   Line "Line_420" at 976,739 size 25x0
      Appearance <- "step_vessel_5"
      Visibility <- "step_vessel_5_proses"
   Line "Line_421" at 748,400 size 25x11
      Appearance <- "step_vessel_4"
      Visibility <- "step_vessel_4_proses"
   Line "Line_422" at 752,412 size 36x78
      Appearance <- "step_vessel_4"
      Visibility <- "step_vessel_4_proses"
   Line "Line_423" at 788,488 size 0x11
      Appearance <- "step_vessel_4"
      Visibility <- "step_vessel_4_proses"
   Line "Line_426" at 767,595 size 21x144
      Appearance <- "step_vessel_4"
      Visibility <- "step_vessel_4_proses"
   Line "Line_427" at 788,579 size 0x19
      Appearance <- "step_vessel_4"
      Visibility <- "step_vessel_4_proses"
   Line "Line_428" at 764,739 size 25x0
      Appearance <- "step_vessel_4"
      Visibility <- "step_vessel_4_proses"
   Line "Line_429" at 536,400 size 25x11
      Appearance <- "step_vessel_3"
   Line "Line_430" at 540,412 size 36x78
      Appearance <- "step_vessel_3"
   Line "Line_431" at 576,488 size 0x11
      Appearance <- "step_vessel_3"
   Line "Line_432" at 748,400 size 25x11
      Appearance <- "step_vessel_4"
   Line "Line_433" at 752,412 size 36x78
      Appearance <- "step_vessel_4"
   Line "Line_434" at 788,488 size 0x11
      Appearance <- "step_vessel_4"
   Line "Line_435" at 960,400 size 25x11
      Appearance <- "step_vessel_5"
   Line "Line_436" at 964,412 size 36x78
      Appearance <- "step_vessel_5"
   Line "Line_437" at 1000,488 size 0x11
      Appearance <- "step_vessel_5"
   Line "Line_438" at 1172,400 size 25x11
      Appearance <- "step_vessel_6"
   Line "Line_439" at 1176,412 size 36x78
      Appearance <- "step_vessel_6"
   Line "Line_440" at 1212,488 size 0x11
      Appearance <- "step_vessel_6"
   Line "Line_441" at 1384,400 size 25x11
      Appearance <- "step_vessel_7"
   Line "Line_442" at 1388,412 size 36x78
      Appearance <- "step_vessel_7"
   Line "Line_443" at 1424,488 size 0x11
      Appearance <- "step_vessel_7"
   Line "Line_450" at 555,595 size 21x144
      Appearance <- "step_vessel_3"
   Line "Line_451" at 576,579 size 0x19
      Appearance <- "step_vessel_3"
   Line "Line_452" at 552,739 size 25x0
      Appearance <- "step_vessel_3"
   Line "Line_453" at 767,595 size 21x144
      Appearance <- "step_vessel_4"
   Line "Line_454" at 788,579 size 0x19
      Appearance <- "step_vessel_4"
   Line "Line_455" at 764,739 size 25x0
      Appearance <- "step_vessel_4"
   Line "Line_457" at 979,595 size 21x144
      Appearance <- "step_vessel_5"
   Line "Line_458" at 1000,579 size 0x19
      Appearance <- "step_vessel_5"
   Line "Line_459" at 976,739 size 25x0
      Appearance <- "step_vessel_5"
   Line "Line_461" at 1191,595 size 21x144
      Appearance <- "step_vessel_6"
   Line "Line_462" at 1212,579 size 0x19
      Appearance <- "step_vessel_6"
   Line "Line_463" at 1188,739 size 25x0
      Appearance <- "step_vessel_6"
   Line "Line_464" at 1403,595 size 21x144
      Appearance <- "step_vessel_7"
   Line "Line_465" at 1424,579 size 0x19
      Appearance <- "step_vessel_7"
   Line "Line_466" at 1400,739 size 25x0
      Appearance <- "step_vessel_7"
   Polygon "Polygon_217" at 123,352 size 58x419
      Appearance <- "ISI TANK 1"
      Visibility <- "ISI TANK 1"
   Line "Line_468" at 124,432 size 57x0
      Visibility <- "ISI TANK 1"
   Line "Line_469" at 142,385 size 21x0
      Visibility <- "ISI TANK 1"
   Line "Line_470" at 124,680 size 56x0
      Visibility <- "ISI TANK 1"
   Polygon "Polygon_218" at 335,352 size 58x419
      Appearance <- "ISI TANK 2"
      Visibility <- "ISI TANK 2"
   Line "Line_471" at 336,432 size 57x0
      Visibility <- "ISI TANK 2"
   Line "Line_472" at 354,385 size 21x0
      Visibility <- "ISI TANK 2"
   Line "Line_473" at 336,680 size 56x0
      Visibility <- "ISI TANK 2"
   Polygon "Polygon_219" at 547,352 size 58x419
      Appearance <- "ISI TANK 3"
      Visibility <- "ISI TANK 3"
   Line "Line_474" at 548,432 size 57x0
      Visibility <- "ISI TANK 3"
   Line "Line_475" at 566,385 size 21x0
      Visibility <- "ISI TANK 3"
   Line "Line_476" at 548,680 size 56x0
      Visibility <- "ISI TANK 3"
   Polygon "Polygon_220" at 759,352 size 58x419
      Appearance <- "ISI TANK 4"
      Visibility <- "ISI TANK 4"
   Line "Line_477" at 760,432 size 57x0
      Visibility <- "ISI TANK 4"
   Line "Line_478" at 778,385 size 21x0
      Visibility <- "ISI TANK 4"
   Line "Line_479" at 760,680 size 56x0
      Visibility <- "ISI TANK 4"
   Polygon "Polygon_221" at 971,352 size 58x419
      Appearance <- "ISI TANK 5"
      Visibility <- "ISI TANK 5"
   Line "Line_480" at 972,432 size 57x0
      Visibility <- "ISI TANK 5"
   Line "Line_481" at 990,385 size 21x0
      Visibility <- "ISI TANK 5"
   Line "Line_482" at 972,680 size 56x0
      Visibility <- "ISI TANK 5"
   Polygon "Polygon_222" at 1183,352 size 58x419
      Appearance <- "ISI TANK 6"
      Visibility <- "ISI TANK 6"
   Line "Line_483" at 1184,432 size 57x0
      Visibility <- "ISI TANK 6"
   Line "Line_484" at 1202,385 size 21x0
      Visibility <- "ISI TANK 6"
   Line "Line_485" at 1184,680 size 56x0
      Visibility <- "ISI TANK 6"
   Polygon "Polygon_223" at 1395,352 size 58x419
      Appearance <- "ISI TANK 7"
      Visibility <- "ISI TANK 7"
   Line "Line_486" at 1396,432 size 57x0
      Visibility <- "ISI TANK 7"
   Line "Line_487" at 1414,385 size 21x0
      Visibility <- "ISI TANK 7"
   Line "Line_488" at 1396,680 size 56x0
      Visibility <- "ISI TANK 7"
   Line "Line_489" at 105,898 size 0x48
      Visibility <- "step_vessel_1_proses"
      Appearance <- "step_vessel_1_proses"
   Line "Line_490" at 102,948 size 40x0
      Appearance <- "step_vessel_1_proses"
      Visibility <- "step_vessel_1_proses"
   Rectangle "Rectangle_10" at 75,874 size 1423x33
      Appearance <- "step_vessel_1_proses"
      Visibility <- "step_vessel_1_proses"
   Line "Line_491" at 105,898 size 0x48
      Appearance <- "step_vessel_2_proses"
      Visibility <- "step_vessel_2_proses"
   Line "Line_492" at 102,948 size 40x0
      Appearance <- "step_vessel_2_proses"
      Visibility <- "step_vessel_2_proses"
   Rectangle "Rectangle_11" at 75,874 size 1423x33
      Visibility <- "step_vessel_2_proses"
      Appearance <- "step_vessel_2_proses"
   Line "Line_493" at 105,898 size 0x48
      Appearance <- "step_vessel_3_proses"
      Visibility <- "step_vessel_3_proses"
   Line "Line_494" at 102,948 size 40x0
      Appearance <- "step_vessel_3_proses"
      Visibility <- "step_vessel_3_proses"
   Rectangle "Rectangle_12" at 75,874 size 1423x33
      Appearance <- "step_vessel_3_proses"
      Visibility <- "step_vessel_3_proses"
   Group "proses_3" at 75,874 size 1423x74
   Line "Line_495" at 105,898 size 0x48
      Appearance <- "step_vessel_4_proses"
      Visibility <- "step_vessel_4_proses"
   Line "Line_496" at 102,948 size 40x0
      Appearance <- "step_vessel_4_proses"
      Visibility <- "step_vessel_4_proses"
   Rectangle "Rectangle_13" at 75,874 size 1423x33
      Appearance <- "step_vessel_4_proses"
      Visibility <- "step_vessel_4_proses"
   Group "proses_4" at 75,874 size 1423x74
   Line "Line_497" at 105,898 size 0x48
      Appearance <- "step_vessel_5_proses"
      Visibility <- "step_vessel_5_proses"
   Line "Line_498" at 102,948 size 40x0
      Appearance <- "step_vessel_5_proses"
      Visibility <- "step_vessel_5_proses"
   Rectangle "Rectangle_14" at 75,874 size 1423x33
      Appearance <- "step_vessel_5_proses"
      Visibility <- "step_vessel_5_proses"
   Group "proses_5" at 75,874 size 1423x74
   Line "Line_499" at 105,898 size 0x48
      Visibility <- "step_vessel_6_proses"
      Appearance <- "step_vessel_6_proses"
   Line "Line_500" at 102,948 size 40x0
      Appearance <- "step_vessel_6_proses"
      Visibility <- "step_vessel_6_proses"
   Rectangle "Rectangle_15" at 75,874 size 1423x33
      Appearance <- "step_vessel_6_proses"
      Visibility <- "step_vessel_6_proses"
   Group "proses_6" at 75,874 size 1423x74
   Line "Line_501" at 105,898 size 0x48
      Visibility <- "step_vessel_7_proses"
      Appearance <- "step_vessel_7_proses"
   Line "Line_502" at 102,948 size 40x0
      Appearance <- "step_vessel_7_proses"
      Visibility <- "step_vessel_7_proses"
   Rectangle "Rectangle_16" at 75,874 size 1423x33
      Visibility <- "step_vessel_7_proses"
      Appearance <- "step_vessel_7_proses"
   Group "proses_7" at 75,874 size 1423x74
   Line "Line_379" at 324,400 size 25x11
      Appearance <- "step_vessel_2"
   Line "Line_380" at 328,412 size 36x78
      Appearance <- "step_vessel_2"
   Line "Line_381" at 364,488 size 0x11
      Appearance <- "step_vessel_2"
   Line "Line_505" at 343,595 size 21x144
      Appearance <- "step_vessel_2"
   Line "Line_506" at 364,579 size 0x19
      Appearance <- "step_vessel_2"
   Line "Line_507" at 340,739 size 25x0
      Appearance <- "step_vessel_2"

screen "storage" 1600x1200
   GraphicView "Graphic view_3" at 191,109 size 312x345; Picture "Graphic_8"
   GraphicView "Graphic view_1" at 191,538 size 312x345; Picture "Graphic_8"
   Group "Group" at 704,26 size 95x303; Picture "Graphic_10"
   Group "Group_2" at 704,453 size 95x303; Picture "Graphic_10"
   Group "Group_3" at 898,453 size 95x303; Picture "Graphic_10"
   Group "Group_4" at 898,26 size 95x303; Picture "Graphic_10"
   GraphicView "Graphic view_45" at 1130,217 size 45x48; Picture "Graphic_56"
   GraphicView "Graphic view_44" at 1130,147 size 47x75; Picture "Graphic_55"
   GraphicView "Graphic view_46" at 1218,217 size 45x48; Picture "Graphic_56"
   GraphicView "Graphic view_47" at 1218,147 size 47x75; Picture "Graphic_55"
   GraphicView "Graphic view_49" at 1130,662 size 45x48; Picture "Graphic_56"
   GraphicView "Graphic view_50" at 1130,592 size 47x75; Picture "Graphic_55"
   GraphicView "Graphic view_51" at 1218,662 size 45x48; Picture "Graphic_56"
   GraphicView "Graphic view_52" at 1218,592 size 47x75; Picture "Graphic_55"
   Button "Button_1" at 633,851 size 192x32; TextOn 'Screen_1'; TextOff 'Vessel'
      on Click: ActivateScreen("vessel", 0)
   Button "Button_2" at 880,851 size 192x32; TextOn 'Screen_3'; TextOff 'Supply'
      on Click: ActivateScreen("supply", 0)
   TextField "Text field_9" at 1484,420 size 16x22; Text 'D'
   IOField "I/O field_25" at 1216,276 size 38x17; FormatPattern 9999999
      Appearance <- "VP FLAVOUR"
   TextField "Text field_13" at 1252,276 size 25x18; Text 'bar'
   IOField "I/O field_26" at 1022,229 size 38x17; FormatPattern 9999999
      Appearance <- "VP FLAVOUR"
   TextField "Text field_14" at 1058,229 size 23x18; Text 'º C'
   IOField "I/O field_1" at 1116,24 size 38x17; FormatPattern 9999999
      Appearance <- "VP FLAVOUR"
   TextField "Text field_10" at 1152,24 size 25x18; Text 'bar'
   IOField "I/O field_2" at 1022,655 size 38x17; FormatPattern 9999999
      Appearance <- "VP HIDROLIC"
   TextField "Text field_1" at 1058,655 size 23x18; Text 'º C'
   IOField "I/O field_3" at 1216,724 size 38x17; FormatPattern 9999999
      Appearance <- "VP HIDROLIC"
   TextField "Text field_5" at 1252,724 size 25x18; Text 'bar'
   IOField "I/O field_4" at 1116,480 size 38x17; FormatPattern 9999999
      Appearance <- "VP HIDROLIC"
   TextField "Text field_4" at 1152,480 size 25x18; Text 'bar'
   IOField "I/O field_5" at 798,711 size 38x17; FormatPattern 9999999
      Appearance <- "VP HIDROLIC"
   TextField "Text field_6" at 834,711 size 23x18; Text 'º C'
   IOField "I/O field_6" at 798,287 size 38x17; FormatPattern 9999999
      Appearance <- "VP FLAVOUR"
   TextField "Text field_7" at 834,287 size 23x18; Text 'º C'
   IOField "I/O field_7" at 614,47 size 38x17; FormatPattern 9999999
      Appearance <- "VP FLAVOUR"
   TextField "Text field_2" at 650,47 size 23x18; Text 'º C'
   IOField "I/O field_8" at 614,471 size 38x17; FormatPattern 9999999
      Appearance <- "VP HIDROLIC"
   TextField "Text field_3" at 650,471 size 23x18; Text 'º C'
   TextField "Text field_8" at 195,529 size 138x23; Text 'TANK HIDROLIK'
   TextField "Text field_12" at 1449,457 size 117x23; Text 'FROM VESSEL'
   GraphicView "Graphic view_4" at 17,916 size 156x94; Picture "Graphic_72"
   GraphicView "Graphic view_7" at 17,481 size 156x94; Picture "Graphic_72"
   Group "Group_10" at 209,458 size 22x12
   Group "Group_1" at 209,890 size 22x12
   Group "Group_6" at 985,57 size 363x395
   Group "Group_8" at 792,83 size 114x184
   Group "Group_11" at 346,86 size 364x39
   Group "Group_12" at 346,86 size 364x39
   Group "Group_13" at 984,507 size 451x318
   Group "Group_15" at 790,516 size 116x179
   Group "Group_17" at 346,513 size 364x42
   Group "Group_18" at 346,513 size 364x42
   Circle "Circle_1" at 320,266 size 43x43
      Appearance <- "tank flavour OK"
   Circle "Circle_2" at 320,698 size 43x43
      Appearance <- "tank hidrolic OK"
   Button "Button_3" at 633,812 size 96x32; TextOff 'Transfer'
      on Press: function_b14e0dd5("transfer", 0)
   Button "Button_4" at 790,810 size 109x34; TextOff 'Auto'; TextList "moded"
      on Click: InvertBit("mode")
      ProcessValue <- "mode"
      Appearance <- "mode"
   Group "Group_19" at 1366,449 size 144x36
   Group "Group_20" at 1366,449 size 144x36
   Group "Group_21" at 1366,449 size 144x36
   Group "Group_22" at 1366,449 size 144x36
   Group "Group_23" at 1366,449 size 144x36
   Group "Group_24" at 1366,449 size 144x36
   Group "Group_25" at 1366,449 size 144x36
   Group "Group_26" at 1366,449 size 144x36
   TextField "Text field_11" at 197,101 size 133x23; Text 'TANK FLAVOUR'
   Button "Button_5" at 17,587 size 96x32; TextOff 'Start'
      on Press: function_b14e0dd5("StartVPpumpFlavour", 0)
   Button "Button_6" at 17,627 size 96x32; TextOff 'Stop'
      on Press: function_b14e0dd5("StopVPpumpFlavour", 0)
   Rectangle "Rectangle_1" at 77,519 size 38x30
      Appearance <- "VP PUMP FLAVOUR"
   Button "Button_7" at 17,1019 size 96x32; TextOff 'Start'
      on Press: function_b14e0dd5("StartVPpumpHidrolic", 0)
   Button "Button_8" at 17,1059 size 96x32; TextOff 'Stop'
      on Press: function_b14e0dd5("StopVPpumpHidrolic", 0)
   Rectangle "Rectangle_2" at 77,951 size 38x30
      Appearance <- "VP PUMP HIDROLIC"
   Group "Group_27" at 156,387 size 190x99
   Group "Group_28" at 156,819 size 190x104
   Group "Group_14" at 984,507 size 451x318
   Button "Button_21" at 1128,851 size 192x32; TextOn 'Screen_3'; TextOff 'EMERGENCY'
      on Click: InvertBit("EMERGENCY")
      Appearance <- "EMERGENCY"
   GraphicView "Graphic view_2" at 704,26 size 95x303; Picture "Graphic_10"
   GraphicView "Graphic view_5" at 704,453 size 95x303; Picture "Graphic_10"
   GraphicView "Graphic view_6" at 898,453 size 95x303; Picture "Graphic_10"
   GraphicView "Graphic view_17" at 898,26 size 95x303; Picture "Graphic_10"
   Line "Line_32" at 156,461 size 0x25
      Appearance <- "VP PUMP FLAVOUR"
   Line "Line_33" at 156,464 size 53x0
      Appearance <- "VP PUMP FLAVOUR"
   Line "Line_34" at 233,464 size 111x0
      Appearance <- "VP PUMP FLAVOUR"
   Line "Line_35" at 346,387 size 0x80
      Appearance <- "VP PUMP FLAVOUR"
   Polygon "Polygon_9" at 209,458 size 11x11
      Appearance <- "VP PUMP FLAVOUR"
   Polygon "Polygon_10" at 220,459 size 11x11
      Appearance <- "VP PUMP FLAVOUR"
   Line "Line_37" at 156,896 size 53x0
      Appearance <- "VP PUMP HIDROLIC"
   Line "Line_36" at 156,893 size 0x30
      Appearance <- "VP PUMP HIDROLIC"
   Line "Line_38" at 233,896 size 111x0
      Appearance <- "VP PUMP HIDROLIC"
   Line "Line_39" at 346,819 size 0x80
      Appearance <- "VP PUMP HIDROLIC"
   Polygon "Polygon_1" at 209,890 size 11x11
      Appearance <- "VP PUMP HIDROLIC"
   Polygon "Polygon_2" at 220,891 size 11x11
      Appearance <- "VP PUMP HIDROLIC"
   Group "Group_5" at 1345,443 size 22x12
   Group "VP HIDROLIC" at 1426,485 size 12x22
   Polygon "Polygon_3" at 1345,443 size 11x11
      Appearance <- "VP FLAVOUR"
   Polygon "Polygon_4" at 1356,444 size 11x11
      Appearance <- "VP FLAVOUR"
   Polygon "Polygon_205" at 1426,496 size 11x11
      Appearance <- "VP HIDROLIC"
   Polygon "Polygon_206" at 1427,485 size 11x11
      Appearance <- "VP HIDROLIC"
   Group "Group_7" at 985,57 size 363x395
   Group "Group_9" at 792,83 size 114x184
   Group "Group_16" at 790,516 size 116x179
   Line "Line_43" at 985,265 size 113x0
      Visibility <- "VP FLAVOUR"
   Line "Line_44" at 1095,58 size 0x208
      Visibility <- "VP FLAVOUR"
   Line "Line_45" at 1092,57 size 111x0
      Visibility <- "VP FLAVOUR"
   Line "Line_46" at 1200,58 size 0x394
      Visibility <- "VP FLAVOUR"
   Line "Line_47" at 1201,449 size 147x0
      Visibility <- "VP FLAVOUR"
   Line "Line_48" at 846,86 size 60x0
      Visibility <- "VP FLAVOUR"
   Line "Line_49" at 847,83 size 0x184
      Visibility <- "VP FLAVOUR"
   Line "Line_50" at 792,265 size 58x0
      Visibility <- "VP FLAVOUR"
   Line "Line_51" at 348,89 size 362x0
      Visibility <- "VP FLAVOUR"
   Line "Line_52" at 346,86 size 0x39
      Visibility <- "VP FLAVOUR"
   Line "Line_58" at 984,692 size 112x0
      Visibility <- "VP HIDROLIC"
   Line "Line_57" at 1095,515 size 0x180
      Visibility <- "VP HIDROLIC"
   Line "Line_56" at 1092,516 size 111x0
      Visibility <- "VP HIDROLIC"
   Line "Line_55" at 1200,517 size 0x308
      Visibility <- "VP HIDROLIC"
   Line "Line_54" at 1202,822 size 233x0
      Visibility <- "VP HIDROLIC"
   Line "Line_53" at 1432,507 size 0x316
      Visibility <- "VP HIDROLIC"
   Line "Line_59" at 844,516 size 62x0
      Visibility <- "VP HIDROLIC"
   Line "Line_60" at 847,518 size 0x177
      Visibility <- "VP HIDROLIC"
   Line "Line_61" at 790,692 size 58x0
      Visibility <- "VP HIDROLIC"
   Line "Line_62" at 347,516 size 363x0
      Visibility <- "VP HIDROLIC"
   Line "Line_63" at 346,513 size 0x42
      Visibility <- "VP HIDROLIC"
   Line "Line_42" at 1366,449 size 144x0
      Visibility <- "VP 13"
   Line "Line_64" at 1432,450 size 0x35
      Visibility <- "VP 13"
   Line "Line_65" at 1366,449 size 144x0
      Visibility <- "VP 22"
   Line "Line_66" at 1432,450 size 0x35
      Visibility <- "VP 22"
   Line "Line_67" at 1366,449 size 144x0
      Visibility <- "VP 34"
   Line "Line_68" at 1432,450 size 0x35
      Visibility <- "VP 34"
   Line "Line_69" at 1366,449 size 144x0
      Visibility <- "VP 46"
   Line "Line_70" at 1432,450 size 0x35
      Visibility <- "VP 46"
   Line "Line_71" at 1366,449 size 144x0
      Visibility <- "VP 58"
   Line "Line_72" at 1432,450 size 0x35
      Visibility <- "VP 58"
   Line "Line_73" at 1366,449 size 144x0
      Visibility <- "VP 70"
   Line "Line_74" at 1432,450 size 0x35
      Visibility <- "VP 70"
   Line "Line_75" at 1366,449 size 144x0
      Visibility <- "VP 82"
   Line "Line_76" at 1432,450 size 0x35
      Visibility <- "VP 82"

screen "supply" 1600x1200
   GraphicView "Graphic view_3" at 234,333 size 290x547; Picture "Graphic_12"
   GraphicView "Graphic view_4" at 619,711 size 89x141; Picture "Graphic_13"
   GraphicView "Graphic view_343" at 847,481 size 118x241; Picture "Graphic_48"
   GraphicView "Graphic view_1" at 1112,481 size 118x241; Picture "Graphic_48"
   Button "Button_1" at 525,950 size 192x32; TextOn 'Screen_1'; TextOff 'VESSEL'
      on Click: ActivateScreen("vessel", 0)
   Button "Button_2" at 745,950 size 192x32; TextOn 'Screen_2'; TextOff 'STORAGE'
      on Click: ActivateScreen("storage", 0)
   Rectangle "Rectangle_5" at 647,745 size 50x66
      Appearance <- "CV AIR 1"
   IOField "I/O field_26" at 976,365 size 38x17; FormatPattern 9999
      ProcessValue <- "temperature THE 1"
      Appearance <- "temperature THE 1"
   TextField "Text field_14" at 1012,365 size 23x18; Text 'º C'
   IOField "I/O field_1" at 829,331 size 38x17; FormatPattern 9999
      ProcessValue <- "pressure steam supply"
      Appearance <- "pressure steam supply"
   TextField "Text field_10" at 865,331 size 25x18; Text 'bar'
   IOField "I/O field_2" at 1272,365 size 38x17; FormatPattern 9999
      ProcessValue <- "temperature THE 2"
      Appearance <- "temperature THE 2"
   TextField "Text field_3" at 1308,365 size 23x18; Text 'º C'
   IOField "I/O field_3" at 852,365 size 38x17; FormatPattern 9999999
   TextField "Text field_1" at 888,365 size 23x18; Text 'º C'
   TextField "Text field_2" at 1392,292 size 15x22; Text 'C'
   TextField "Text field_4" at 1393,395 size 15x22; Text 'B'
   TextField "Text field_12" at 1421,340 size 93x23; Text 'TO VESSEL'
   Group "Group_16" at 803,389 size 22x12
   Group "Group" at 789,293 size 14x259
   Group "Group_1" at 803,546 size 22x12
   Group "Group_2" at 1067,389 size 22x12
   Group "Group_4" at 1054,291 size 14x263
   Group "Group_3" at 1067,546 size 22x12
   Button "Button_5" at 88,467 size 109x34; TextOff 'Supply'
      on Press: function_b14e0dd5("supply", 0)
   Button "Button_3" at 88,520 size 109x34; TextOff 'Auto'; TextList "moded"
      on Click: InvertBit("mode")
      ProcessValue <- "mode"
      Appearance <- "mode"
   Button "Button_21" at 966,950 size 192x32; TextOn 'Screen_3'; TextOff 'EMERGENCY'
      on Click: InvertBit("EMERGENCY")
      Appearance <- "EMERGENCY"
   Polygon "Polygon_21" at 803,389 size 11x11
      Appearance <- "CV AIR 1"
   Polygon "Polygon_22" at 814,390 size 11x11
      Appearance <- "CV AIR 1"
   Polygon "Polygon_1" at 803,546 size 11x11
      Appearance <- "CV STEAM 1"
   Polygon "Polygon_2" at 814,547 size 11x11
      Appearance <- "CV STEAM 1"
   Polygon "Polygon_3" at 1067,389 size 11x11
      Appearance <- "CV AIR 2"
   Polygon "Polygon_4" at 1078,390 size 11x11
      Appearance <- "CV AIR 2"
   Polygon "Polygon_5" at 1067,546 size 11x11
      Appearance <- "CV STEAM 2"
   Polygon "Polygon_6" at 1078,547 size 11x11
      Appearance <- "CV STEAM 2"

screen "Screen_4" 1600x1200
   GraphicView "Graphic view_36" at 284,492 size 63x442; Picture "Graphic_1"
   Group "Group" at 376,500 size 58x419

Template "Template_1" 1600x1200
   GraphicView "Graphic view_1" at 0,6 size 1590x1184; Picture "machine simulation"

VB script "Vessel1"
   If SmartTags("step_vessel_1")<>0 Then
   	If SmartTags("VB 1") = True Then
   		SmartTags("pipa bawah") = 10
   	End If
   Else
   	b21d3eaf-4e31-425c-ad1a-ba4e4002cacc pipa bawah,0 		
   End If

VB script "Vessel2"
   If SmartTags("step_vessel_2")<>0 Then
   	If SmartTags("VB 2") = True Then
   		b21d3eaf-4e31-425c-ad1a-ba4e4002cacc pipa bawah,10	
   	End If
   Else
   	b21d3eaf-4e31-425c-ad1a-ba4e4002cacc pipa bawah,0 	
   End If

VB script "Vessel3"
   If SmartTags("step_vessel_3")<>0 Then
   	If SmartTags("VB 3") = True Then
   		SmartTags("pipa bawah") = 10
   	End If
   Else
   	SmartTags("pipa bawah") = 0	
   End If

VB script "Vessel4"
   If SmartTags("step_vessel_4")<>0 Then
   	If SmartTags("VB 4") = True Then
   		SmartTags("pipa bawah") = 10
   	End If
   Else
   	SmartTags("pipa bawah") = 0	
   End If

VB script "Vessel5"
   If SmartTags("step_vessel_5")<>0 Then
   	If SmartTags("VB 5") = True Then
   		SmartTags("pipa bawah") = 10
   	End If
   Else
   	SmartTags("pipa bawah") = 0	
   End If

VB script "Vessel6"
   If SmartTags("step_vessel_6")<>0 Then
   	If SmartTags("VB 6") = True Then
   		SmartTags("pipa bawah") = 10
   	End If
   Else
   	b21d3eaf-4e31-425c-ad1a-ba4e4002cacc pipa bawah,0 	
   End If

VB script "Vessel7"
   If SmartTags("step_vessel_7")<>0 Then
   	If SmartTags("VB 7") = True Then
   		SmartTags("pipa bawah") = 10
   	End If
   Else
   	SmartTags("pipa bawah") = 0	
   End If

VB script "tank"
   If SmartTags("step_isi") = 1 Then 
   	SmartTags("tank 1") = 10
   end if
*)